// TIA Portal project "Delta_Praktika_3" (V17)

(* hardware
DEVICE "S7-1500/ET200MP station_1"  S7-1500 station
   slot 0: "Rail_0"  Rack  6ES7 590-1***0-0AA0
   slot 1: "PLC_2"  CPU 1517TF-3 PN/DP  6ES7 517-3UP00-0AB0  V2.9
      slot 3: "CPU display_1"  6ES7591-1BA00-0AA0
      slot 32768: "PROFINET interface_1"  X1
      slot 33024: "PROFINET interface_2"  X2
      slot 33280: "DP interface_1"  X3
      slot 34817: "Virtual CP interface port_1"  Virtual CP interface port  Virtual CP interface port
DEVICE "ET 200SP station_1"  ET 200SP-Station
   slot 0: "Rack_0"  Rack  6ES5 710-8MAx1
   slot 0: "et200sp"  IM 155-6 PN/2 HF  6ES7 155-6AU01-0CN0  V4.2
   slot 1: "DI 8x24VDC HF_1"  DI 8x24VDC HF  6ES7 131-6BF00-0CA0  V2.0
      slot 1: "DI 8x24VDC HF_1"  DI 8x24VDC HF
   slot 2: "DQ 8x24VDC/0.5A HF_1"  DQ 8x24VDC/0.5A HF  6ES7 132-6BF00-0CA0  V2.0
      slot 1: "DQ 8x24VDC/0.5A HF_1"  DQ 8x24VDC/0.5A HF
   slot 3: "CM 4xIO-Link_1"  CM 4xIO-Link  6ES7 137-6BD00-0BA0  V2.2
      slot 1: "CM 4xIO-Link_1"  6ES7 137-6BD00-0BA0
   slot 4: "Server module_1"  Server module  6ES7 193-6PA00-0AA0  V1.1
      slot 1: "Server module_1"  Server module
   slot 127: "BA 2xRJ45"  BA 2xRJ45  6ES7 193-6AR00-0AA0  V0.0
      slot 1: "Port_1"  X1 P1 R  6ES7 193-6AR00-0AA0  V0.0
      slot 2: "Port_2"  X1 P2 R  6ES7 193-6AR00-0AA0  V0.0
DEVICE "SINAMICS V_1"  SINAMICS V
   slot 0: "SINAMICS V90 PN Rack"  Rail  1.0
   slot 0: "a1"  V90 PN  6SL3 210-5FB10-4UFx  V1.4
      slot 1: "Drive object"  Drive Object
         slot 1: "Module access point"  Module Access Point
         slot 2: "Without PROFIsafe"  No ProfiSafe
         slot 3: "Telegram"  SIEMENS Telegramm 105
DEVICE "SINAMICS V_2"  SINAMICS V
   slot 0: "SINAMICS V90 PN Rack"  Rail  1.0
   slot 0: "a3"  V90 PN  6SL3 210-5FB10-4UFx  V1.4
      slot 1: "Drive object"  Drive Object
         slot 1: "Module access point"  Module Access Point
         slot 2: "Without PROFIsafe"  No ProfiSafe
         slot 3: "Telegram"  SIEMENS Telegramm 105
DEVICE "SINAMICS V_3"  SINAMICS V
   slot 0: "SINAMICS V90 PN Rack"  Rail  1.0
   slot 0: "a2"  V90 PN  6SL3 210-5FB10-4UFx  V1.4
      slot 1: "Drive object"  Drive Object
         slot 1: "Module access point"  Module Access Point
         slot 2: "Without PROFIsafe"  No ProfiSafe
         slot 3: "Telegram"  SIEMENS Telegramm 105
DEVICE "HMI_1"  KTP1200 Basic PN
   slot 0: "HMI_1"  KTP1200 Basic PN  6AV2 123-2MB03-0AX0  17.0.0.0
   slot 1: "HMI_RT_1"  KTP1200 Basic PN  6AV2 123-2MB03-0AX0  17.0.0.0
   slot 5: "HMI_1.IE_CP_1"  PROFINET Interface  17.0.0.0
      slot 1: "Interfaz PROFINET_1"  PROFINET Interface
         slot 1: "Port_1"  Port
*)

// ===== PLC "PLC_2"  CPU 1517TF-3 PN/DP =====
// protected blocks, not shown: "Main_Safety_RTG1", "Main_Safety_RTG1_DB"

VAR_GLOBAL   // PLC tag table "Default tag table"
   "A1_Actor_Interface_AddressIn" AT %I0.0 : "PD_TEL3_IN";
   "A1_Actor_Interface_AddressOut" AT %Q0.0 : "PD_TEL3_OUT";
   "A2_Actor_Interface_AddressIn" AT %I18.0 : "PD_TEL3_IN";
   "A2_Actor_Interface_AddressOut" AT %Q10.0 : "PD_TEL3_OUT";
   "A3_Actor_Interface_AddressIn" AT %I36.0 : "PD_TEL3_IN";
   "A3_Actor_Interface_AddressOut" AT %Q20.0 : "PD_TEL3_OUT";
   "A1_axis_Actor_Interface_AddressIn" AT %I0.0 : "PD_TEL105_IN";
   "A1_axis_Actor_Interface_AddressOut" AT %Q0.0 : "PD_TEL105_OUT";
   "a2_axis_Actor_Interface_AddressIn" AT %I20.0 : "PD_TEL105_IN";
   "a2_axis_Actor_Interface_AddressOut" AT %Q63.0 : "PD_TEL105_OUT";
   "a3_asix_Actor_Interface_AddressIn" AT %I87.0 : "PD_TEL105_IN";
   "a3_asix_Actor_Interface_AddressOut" AT %Q83.0 : "PD_TEL105_OUT";
   "Freno_a1" AT %Q30.1 : Bool;
   "marka_Freno_a1" AT %M30.1 : Bool;
   "marka_Freno_a2" AT %M30.2 : Bool;
   "Freno_a2" AT %Q30.2 : Bool;
   "Freno_a3" AT %Q30.0 : Bool;
   "marka_Freno_a3" AT %M30.0 : Bool;
   "System_Byte" AT %MB256 : Byte;
   "FirstScan" AT %M256.0 : Bool;
   "DiagStatusUpdate" AT %M256.1 : Bool;
   "AlwaysTRUE" AT %M256.2 : Bool;
   "AlwaysFALSE" AT %M256.3 : Bool;
   "Clock_Byte" AT %MB255 : Byte;
   "Clock_10Hz" AT %M255.0 : Bool;
   "Clock_5Hz" AT %M255.1 : Bool;
   "Clock_2.5Hz" AT %M255.2 : Bool;
   "Clock_2Hz" AT %M255.3 : Bool;
   "Clock_1.25Hz" AT %M255.4 : Bool;
   "Clock_1Hz" AT %M255.5 : Bool;
   "Clock_0.625Hz" AT %M255.6 : Bool;
   "Clock_0.5Hz" AT %M255.7 : Bool;
   "Tag_1" AT %M401.0 : Bool;
END_VAR

DATA_BLOCK "Power_DB"   // DB9
{ S7_Optimized_Access := 'TRUE' }
VERSION : 0.1
// stored: InstanceOfName Power
"Power"
BEGIN
END_DATA_BLOCK

DATA_BLOCK "Parametroak"   // DB11
{ S7_Optimized_Access := 'TRUE' }
VERSION : 0.1
   VAR
      Abiadura : LReal := 2.0;
      Azelerazioa : LReal := 40.0;
      Desazelerazioa : LReal := 40.0;
      Jerk : LReal := 400.0;
   END_VAR
BEGIN
END_DATA_BLOCK

DATA_BLOCK "Jog_DB"   // DB14
{ S7_Optimized_Access := 'TRUE' }
VERSION : 0.1
// stored: InstanceOfName Jog
"Jog"
BEGIN
END_DATA_BLOCK

DATA_BLOCK "Hominga_DB"   // DB18
{ S7_Optimized_Access := 'TRUE' }
VERSION : 0.1
// stored: InstanceOfName Hominga
"Hominga"
BEGIN
END_DATA_BLOCK

DATA_BLOCK "Puntuak"   // DB24
{ S7_Optimized_Access := 'TRUE' }
VERSION : 0.1
   VAR
      Puntu_abs_home : Array[1..4] of LReal;
      Puntu_abs_1 : Array[1..4] of LReal;
      Puntu_abs_2 : Array[1..4] of LReal;
      Puntu_rel_1 : Array[1..4] of LReal;
      Puntu_aux_1 : Array[1..3] of LReal;
      Puntu_zirkular_1 : Array[1..4] of LReal;
      HMI_erlatibo_lineal : Array[1..4] of LReal;
      HMI_abs_lineal : Array[1..4] of LReal;
      HMI_abs_zirkular_aux : Array[1..3] of LReal;
      HMI_abs_zirkular_endpoint : Array[1..4] of LReal;
      HMI_abs_ptp : Array[1..4] of LReal;
   END_VAR
BEGIN
   Puntu_abs_home[1] := 0.0;
   Puntu_abs_home[2] := 0.0;
   Puntu_abs_home[3] := -722.59;
   Puntu_abs_home[4] := 0.0;
   Puntu_abs_1[1] := 0.0;
   Puntu_abs_1[2] := 0.0;
   Puntu_abs_1[3] := -700.0;
   Puntu_abs_1[4] := 0.0;
   Puntu_rel_1[1] := 50.0;
   Puntu_rel_1[2] := 0.0;
   Puntu_rel_1[3] := 0.0;
   Puntu_abs_2[1] := 50.0;
   Puntu_abs_2[2] := 50.0;
   Puntu_abs_2[3] := -700.0;
   Puntu_abs_2[4] := 0.0;
   Puntu_aux_1[1] := 50.0;
   Puntu_aux_1[2] := 0.0;
   Puntu_aux_1[3] := -700.0;
   Puntu_zirkular_1[1] := 100.0;
   Puntu_zirkular_1[2] := 0.0;
   Puntu_zirkular_1[3] := -700.0;
   Puntu_zirkular_1[4] := 0.0;
END_DATA_BLOCK

DATA_BLOCK "ParametroakII"   // DB25
{ S7_Optimized_Access := 'TRUE' }
VERSION : 0.1
   VAR
      abiadura : LReal := 10.0;
      azelerazioa : LReal := 20.0;
      desazelerazioa : LReal := 20.0;
      jerk : LReal := 40.0;
   END_VAR
BEGIN
END_DATA_BLOCK

DATA_BLOCK "a1_asix"   // DB2, Motion_DB
{ S7_Optimized_Access := 'TRUE' }
AUTHOR : SIMATIC
FAMILY : MC_1500
VERSION : 6.0
// stored: InstanceOfName TO_PositioningAxis
"TO_PositioningAxis"
BEGIN
END_DATA_BLOCK

DATA_BLOCK "a2_axis"   // DB3, Motion_DB
{ S7_Optimized_Access := 'TRUE' }
AUTHOR : SIMATIC
FAMILY : MC_1500
VERSION : 6.0
// stored: InstanceOfName TO_PositioningAxis
"TO_PositioningAxis"
BEGIN
END_DATA_BLOCK

DATA_BLOCK "a3_axis"   // DB4, Motion_DB
{ S7_Optimized_Access := 'TRUE' }
AUTHOR : SIMATIC
FAMILY : MC_1500
VERSION : 6.0
// stored: InstanceOfName TO_PositioningAxis
"TO_PositioningAxis"
BEGIN
END_DATA_BLOCK

DATA_BLOCK "Delta_Robota"   // DB7, Motion_DB
{ S7_Optimized_Access := 'TRUE' }
AUTHOR : SIMATIC
FAMILY : MC_1500
VERSION : 6.0
// stored: InstanceOfName TO_Kinematics
"TO_Kinematics"
BEGIN
END_DATA_BLOCK

FUNCTION_BLOCK "Power"   // FB2, LAD
{ S7_Optimized_Access := 'TRUE' }
VERSION : 0.1
   VAR_INPUT
      Power_a1 : Bool;
      Power_a2 : Bool;
      Power_a3 : Bool;
   END_VAR
   VAR_OUTPUT
      Status_a1 : Bool;
      Status_a2 : Bool;
      Status_a3 : Bool;
      Error_a1 : Bool;
      Error_a2 : Bool;
      Error_a3 : Bool;
   END_VAR
BEGIN

REGION Network 1
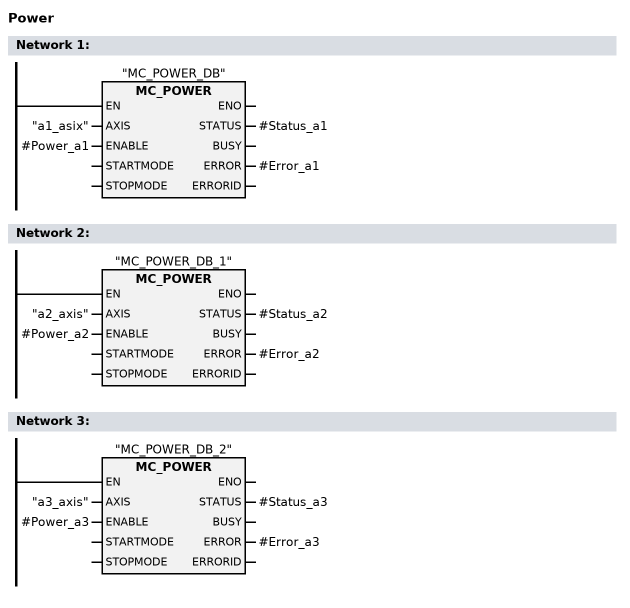
   "MC_POWER_DB"(Axis := "a1_asix", Enable := #Power_a1, Status => #Status_a1, Error => #Error_a1);   // MC_POWER
END_REGION

REGION Network 2
   "MC_POWER_DB_1"(Axis := "a2_axis", Enable := #Power_a2, Status => #Status_a2, Error => #Error_a2);   // MC_POWER
END_REGION

REGION Network 3
   "MC_POWER_DB_2"(Axis := "a3_axis", Enable := #Power_a3, Status => #Status_a3, Error => #Error_a3);   // MC_POWER
END_REGION
END_FUNCTION_BLOCK

FUNCTION_BLOCK "Jog"   // FB3, LAD
{ S7_Optimized_Access := 'TRUE' }
VERSION : 0.1
   VAR_INPUT
      "A1+" : Bool;
      "A1-" : Bool;
      "A2+" : Bool;
      "A2-" : Bool;
      "A3+" : Bool;
      "A3-" : Bool;
   END_VAR
BEGIN

REGION Network 1
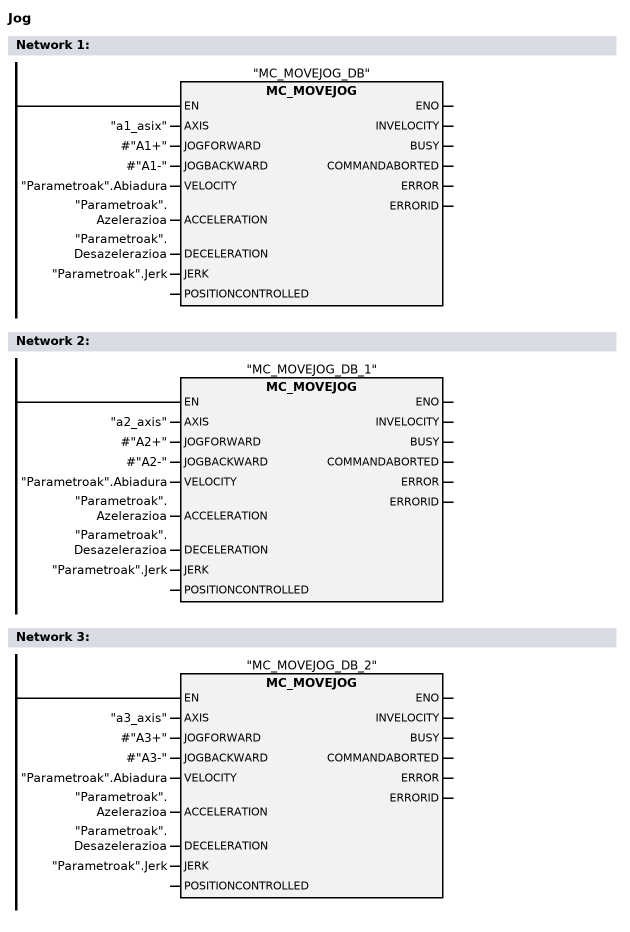
   "MC_MOVEJOG_DB"(Axis := "a1_asix",   // MC_MOVEJOG
                   JogForward := #"A1+",
                   JogBackward := #"A1-",
                   Velocity := "Parametroak".Abiadura,
                   Acceleration := "Parametroak".Azelerazioa,
                   Deceleration := "Parametroak".Desazelerazioa,
                   Jerk := "Parametroak".Jerk);
END_REGION

REGION Network 2
   "MC_MOVEJOG_DB_1"(Axis := "a2_axis",   // MC_MOVEJOG
                     JogForward := #"A2+",
                     JogBackward := #"A2-",
                     Velocity := "Parametroak".Abiadura,
                     Acceleration := "Parametroak".Azelerazioa,
                     Deceleration := "Parametroak".Desazelerazioa,
                     Jerk := "Parametroak".Jerk);
END_REGION

REGION Network 3
   "MC_MOVEJOG_DB_2"(Axis := "a3_axis",   // MC_MOVEJOG
                     JogForward := #"A3+",
                     JogBackward := #"A3-",
                     Velocity := "Parametroak".Abiadura,
                     Acceleration := "Parametroak".Azelerazioa,
                     Deceleration := "Parametroak".Desazelerazioa,
                     Jerk := "Parametroak".Jerk);
END_REGION
END_FUNCTION_BLOCK

FUNCTION_BLOCK "Hominga"   // FB4, LAD
{ S7_Optimized_Access := 'TRUE' }
VERSION : 0.1
   VAR_INPUT
      homing_a1 : Bool;
      homing_a2 : Bool;
      homing_a3 : Bool;
   END_VAR
   VAR_OUTPUT
      Done_a1 : Bool;
      Done_a2 : Bool;
      Done_a3 : Bool;
   END_VAR
BEGIN

REGION Network 1
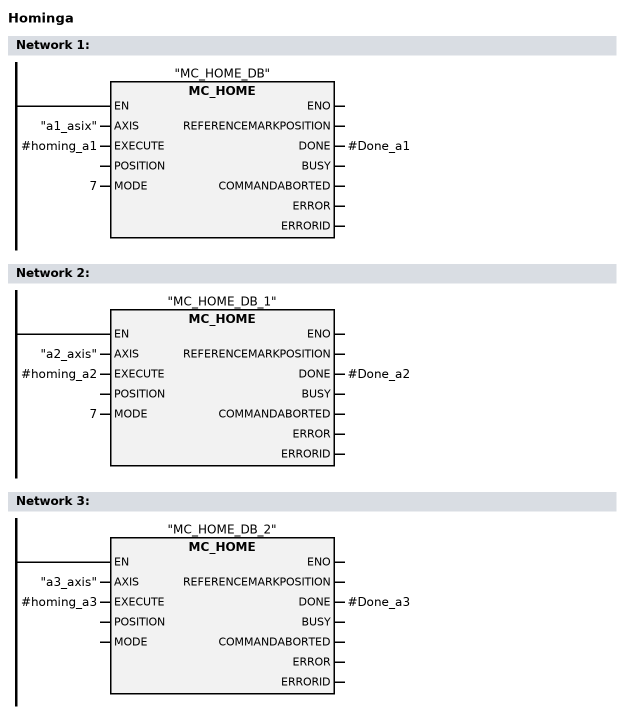
   "MC_HOME_DB"(Axis := "a1_asix", Execute := #homing_a1, Mode := 7, Done => #Done_a1);   // MC_HOME
END_REGION

REGION Network 2
   "MC_HOME_DB_1"(Axis := "a2_axis", Execute := #homing_a2, Mode := 7, Done => #Done_a2);   // MC_HOME
END_REGION

REGION Network 3
   "MC_HOME_DB_2"(Axis := "a3_axis", Execute := #homing_a3, Done => #Done_a3);   // MC_HOME
END_REGION
END_FUNCTION_BLOCK

ORGANIZATION_BLOCK "Main"   // OB1, LAD, ProgramCycle
TITLE = "Main Program Sweep (Cycle)"
{ S7_Optimized_Access := 'TRUE' }
VERSION : 0.1
   VAR_INPUT
      Initial_Call : Bool;   // Initial call of this OB
      Remanence : Bool;   // =True, if remanent data are available
   END_VAR
BEGIN

REGION Network 1
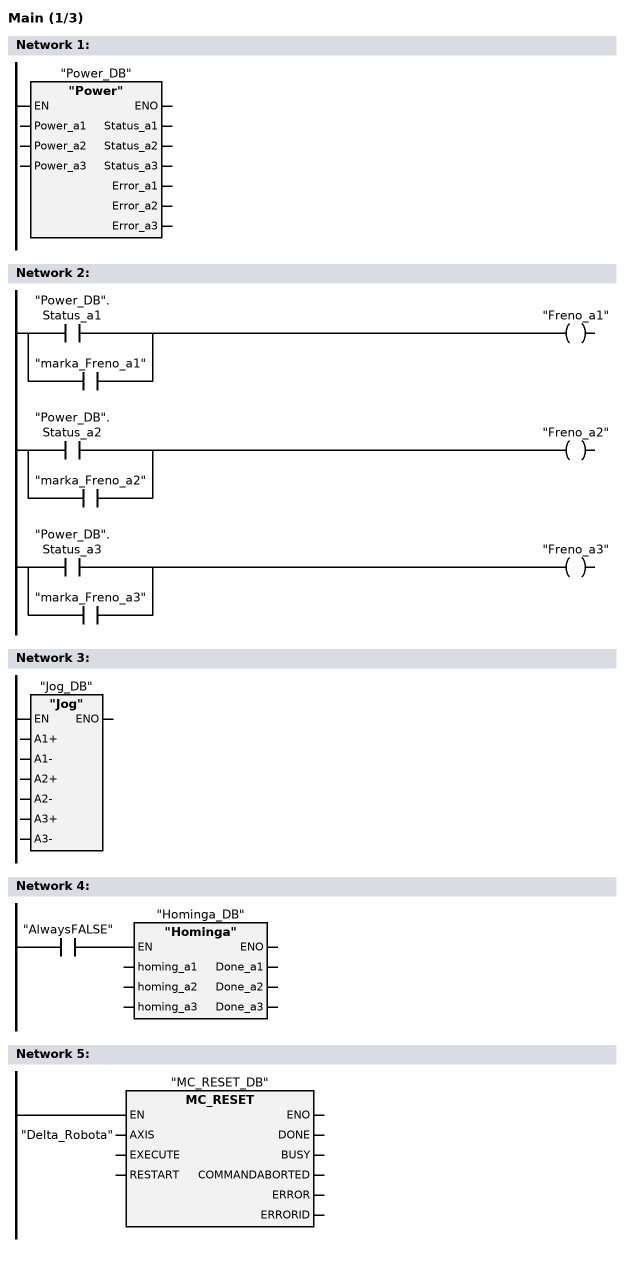
   RUNG wire#powerrail
      "Power_DB"(Power_a1 :=, Power_a2 :=, Power_a3 :=, Status_a1 =>, Status_a2 =>, Status_a3 =>, Error_a1 =>, Error_a2 =>, Error_a3 =>)
   END_RUNG
   // the same network as SCL:
   "Power_DB"();   // "Power"
END_REGION

REGION Network 2
   RUNG wire#powerrail
      Contact( "Power_DB".Status_a1 )
      wire#w1
      Coil( "Freno_a1" )
   END_RUNG
   RUNG wire#powerrail
      Contact( "marka_Freno_a1" )
   END_RUNG wire#w1
   RUNG wire#powerrail
      Contact( "Power_DB".Status_a2 )
      wire#w2
      Coil( "Freno_a2" )
   END_RUNG
   RUNG wire#powerrail
      Contact( "marka_Freno_a2" )
   END_RUNG wire#w2
   RUNG wire#powerrail
      Contact( "Power_DB".Status_a3 )
      wire#w3
      Coil( "Freno_a3" )
   END_RUNG
   RUNG wire#powerrail
      Contact( "marka_Freno_a3" )
   END_RUNG wire#w3
   // the same network as SCL:
   "Freno_a1" := "Power_DB".Status_a1 OR "marka_Freno_a1";
   "Freno_a2" := "Power_DB".Status_a2 OR "marka_Freno_a2";
   "Freno_a3" := "Power_DB".Status_a3 OR "marka_Freno_a3";
END_REGION

REGION Network 3
   RUNG wire#powerrail
      "Jog_DB"("A1+" :=, "A1-" :=, "A2+" :=, "A2-" :=, "A3+" :=, "A3-" :=)
   END_RUNG
   // the same network as SCL:
   "Jog_DB"();   // "Jog"
END_REGION

REGION Network 4
   RUNG wire#powerrail
      Contact( "AlwaysFALSE" )
      "Hominga_DB"(homing_a1 :=, homing_a2 :=, homing_a3 :=, Done_a1 =>, Done_a2 =>, Done_a3 =>)
   END_RUNG
   // the same network as SCL:
   IF "AlwaysFALSE" THEN
       "Hominga_DB"();   // "Hominga"
   END_IF;
END_REGION

REGION Network 5
   "MC_RESET_DB"(Axis := "Delta_Robota");   // MC_RESET
END_REGION

REGION Network 6
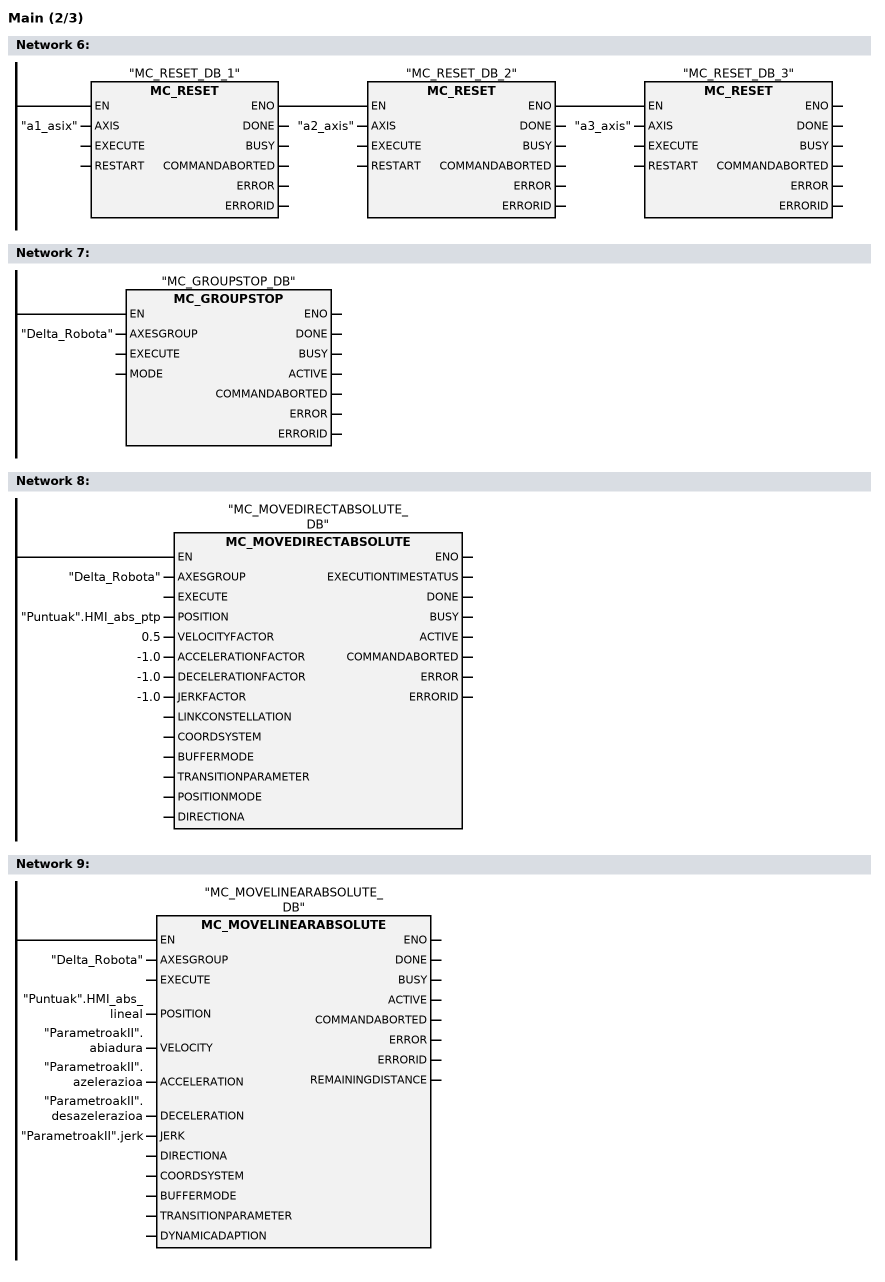
   // ENO of a box is taken as its EN; it also drops when the box reports an error
   "MC_RESET_DB_1"(Axis := "a1_asix");   // MC_RESET
   "MC_RESET_DB_2"(Axis := "a2_axis");   // MC_RESET
   "MC_RESET_DB_3"(Axis := "a3_axis");   // MC_RESET
END_REGION

REGION Network 7
   "MC_GROUPSTOP_DB"(AxesGroup := "Delta_Robota");   // MC_GROUPSTOP
END_REGION

REGION Network 8
   "MC_MOVEDIRECTABSOLUTE_DB"(AxesGroup := "Delta_Robota",   // MC_MOVEDIRECTABSOLUTE
                           Position := "Puntuak".HMI_abs_ptp,
                           VelocityFactor := 0.5,
                           AccelerationFactor := -1.0,
                           DecelerationFactor := -1.0,
                           JerkFactor := -1.0);
END_REGION

REGION Network 9
   "MC_MOVELINEARABSOLUTE_DB"(AxesGroup := "Delta_Robota",   // MC_MOVELINEARABSOLUTE
                           Position := "Puntuak".HMI_abs_lineal,
                           Velocity := "ParametroakII".abiadura,
                           Acceleration := "ParametroakII".azelerazioa,
                           Deceleration := "ParametroakII".desazelerazioa,
                           Jerk := "ParametroakII".jerk);
END_REGION

REGION Network 10
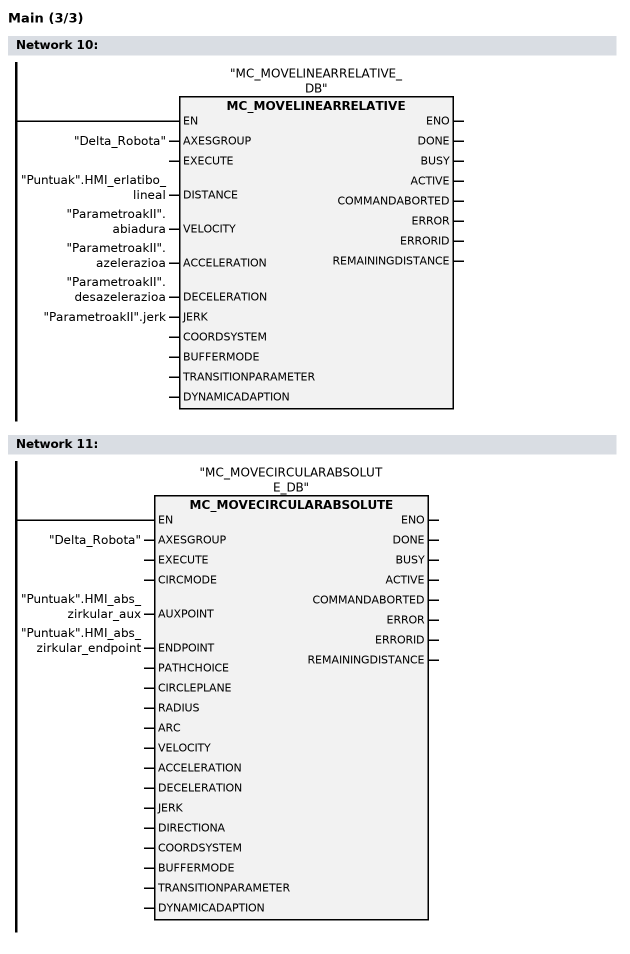
   "MC_MOVELINEARRELATIVE_DB"(AxesGroup := "Delta_Robota",   // MC_MOVELINEARRELATIVE
                           Distance := "Puntuak".HMI_erlatibo_lineal,
                           Velocity := "ParametroakII".abiadura,
                           Acceleration := "ParametroakII".azelerazioa,
                           Deceleration := "ParametroakII".desazelerazioa,
                           Jerk := "ParametroakII".jerk);
END_REGION

REGION Network 11
   "MC_MOVECIRCULARABSOLUTE_DB"(AxesGroup := "Delta_Robota",   // MC_MOVECIRCULARABSOLUTE
                           AuxPoint := "Puntuak".HMI_abs_zirkular_aux,
                           EndPoint := "Puntuak".HMI_abs_zirkular_endpoint);
END_REGION
END_ORGANIZATION_BLOCK

(* ===== HMI "HMI_RT_1" =====
system functions are stored by id; their names below are inferred from use
connection "HMI_Conexión_2": ETHERNET, SMART_S7_1500_OMS

HMI tags "Tabla de variables estándar"
   "Delta_Robota_TcpInWcs_x_Position" : LReal = PLC Delta_Robota.TcpInWcs.x.Position, 1 s
   "Power_DB_Power_a1" : Bool = PLC Power_DB.Power_a1, 1 s
   "Jog_DB_A1+" : Bool = PLC Jog_DB.A1+, 1 s
   "a1_asix_ActualPosition" : LReal = PLC a1_asix.ActualPosition, 1 s
   "Power_DB_Power_a2" : Bool = PLC Power_DB.Power_a2, 1 s
   "Power_DB_Power_a3" : Bool = PLC Power_DB.Power_a3, 1 s
   "Tag_2" : Bool = PLC marka_Freno_a1 AT %M30.1, 1 s
   "Tag_3" : Bool = PLC marka_Freno_a2 AT %M30.2, 1 s
   "Tag_6" : Bool = PLC marka_Freno_a3 AT %M30.0, 1 s
   "Jog_DB_A1-" : Bool = PLC Jog_DB.A1-, 1 s
   "Jog_DB_A2+" : Bool = PLC Jog_DB.A2+, 1 s
   "Jog_DB_A2-" : Bool = PLC Jog_DB.A2-, 1 s
   "Jog_DB_A3+" : Bool = PLC Jog_DB.A3+, 1 s
   "Jog_DB_A3-" : Bool = PLC Jog_DB.A3-, 1 s
   "Tag_1" : Bool = PLC Freno_a1 AT %Q30.1, 1 s
   "Tag_4" : Bool = PLC Freno_a2 AT %Q30.2, 1 s
   "a3_axis_ActualPosition" : LReal = PLC a3_axis.ActualPosition, 1 s
   "Tag_5" : Bool = PLC Freno_a3 AT %Q30.0, 1 s
   "Delta_Robota_TcpInWcs_y_Position" : LReal = PLC Delta_Robota.TcpInWcs.y.Position, 1 s
   "Delta_Robota_TcpInWcs_z_Position" : LReal = PLC Delta_Robota.TcpInWcs.z.Position, 1 s
   "a2_axis_ActualPosition" : LReal = PLC a2_axis.ActualPosition, 1 s
   "MC_GROUPSTOP_DB_Execute" : Bool = PLC MC_GROUPSTOP_DB.Execute, 1 s
   "MC_RESET_DB_Execute" : Bool = PLC MC_RESET_DB.Execute, 1 s
   "Puntuak_HMI_erlatibo_lineal{1}" : LReal = PLC Puntuak.HMI_erlatibo_lineal[1], 1 s
   "Puntuak_HMI_erlatibo_lineal{2}" : LReal = PLC Puntuak.HMI_erlatibo_lineal[2], 1 s
   "Puntuak_HMI_erlatibo_lineal{3}" : LReal = PLC Puntuak.HMI_erlatibo_lineal[3], 1 s
   "Puntuak_HMI_abs_lineal{1}" : LReal = PLC Puntuak.HMI_abs_lineal[1], 1 s
   "Puntuak_HMI_abs_lineal{2}" : LReal = PLC Puntuak.HMI_abs_lineal[2], 1 s
   "Puntuak_HMI_abs_lineal{3}" : LReal = PLC Puntuak.HMI_abs_lineal[3], 1 s
   "Puntuak_HMI_abs_ptp{1}" : LReal = PLC Puntuak.HMI_abs_ptp[1], 1 s
   "Puntuak_HMI_abs_ptp{2}" : LReal = PLC Puntuak.HMI_abs_ptp[2], 1 s
   "Puntuak_HMI_abs_ptp{3}" : LReal = PLC Puntuak.HMI_abs_ptp[3], 1 s
   "MC_MOVELINEARABSOLUTE_DB_Execute" : Bool = PLC MC_MOVELINEARABSOLUTE_DB.Execute, 1 s
   "MC_MOVEDIRECTABSOLUTE_DB_Execute" : Bool = PLC MC_MOVEDIRECTABSOLUTE_DB.Execute, 1 s
   "MC_MOVELINEARRELATIVE_DB_Execute" : Bool = PLC MC_MOVELINEARRELATIVE_DB.Execute, 1 s
   "Puntuak_HMI_abs_zirkular_aux{1}" : LReal = PLC Puntuak.HMI_abs_zirkular_aux[1], 1 s
   "Puntuak_HMI_abs_zirkular_aux{2}" : LReal = PLC Puntuak.HMI_abs_zirkular_aux[2], 1 s
   "Puntuak_HMI_abs_zirkular_aux{3}" : LReal = PLC Puntuak.HMI_abs_zirkular_aux[3], 1 s
   "Puntuak_HMI_abs_zirkular_endpoint{1}" : LReal = PLC Puntuak.HMI_abs_zirkular_endpoint[1], 1 s
   "Puntuak_HMI_abs_zirkular_endpoint{2}" : LReal = PLC Puntuak.HMI_abs_zirkular_endpoint[2], 1 s
   "Puntuak_HMI_abs_zirkular_endpoint{3}" : LReal = PLC Puntuak.HMI_abs_zirkular_endpoint[3], 1 s
   "MC_MOVECIRCULARABSOLUTE_DB_Execute" : Bool = PLC MC_MOVECIRCULARABSOLUTE_DB.Execute, 1 s

screen "Imagen_1" 1280x800
   Button "Botón_1" at 38,159 size 96x32; TextOff 'A1+'
      on Press: function_b14e0dd5("Jog_DB_A1+", 0)
   Button "Botón_2" at 175,159 size 96x32; TextOff 'A1-'
      on Press: function_b14e0dd5("Jog_DB_A1-", 0)
   Button "Botón_3" at 40,207 size 96x32; TextOff 'A2+'
      on Press: function_b14e0dd5("Jog_DB_A2+", 0)
   Button "Botón_4" at 175,207 size 96x32; TextOff 'A2-'
      on Press: function_b14e0dd5("Jog_DB_A2-", 0)
   Button "Botón_5" at 40,255 size 96x32; TextOff 'A3+'
      on Press: function_b14e0dd5("Jog_DB_A3+", 0)
   Button "Botón_6" at 175,255 size 96x32; TextOff 'A3-'
      on Press: function_b14e0dd5("Jog_DB_A3-", 0)
   Button "Botón_10" at 926,70 size 96x32; TextOff 'Stop'
      on Press: function_b14e0dd5("MC_GROUPSTOP_DB_Execute", 0)
   Button "Botón_11" at 1061,70 size 96x32; TextOff 'Reset'
      on Press: function_b14e0dd5("MC_RESET_DB_Execute", 0)
   TextField "Campo de texto_1" at 68,12 size 306x23; Text 'OBJETO TEKNOLOGIKOA BANAKA'
   TextField "Campo de texto_2" at 850,14 size 146x23; Text 'DELTA ROBOTA'
   Circle "Círculo_1" at 415,164 size 19x19
      Appearance <- "Tag_1"
   Circle "Círculo_2" at 415,212 size 19x19
      Appearance <- "Tag_4"
   Circle "Círculo_3" at 415,260 size 19x19
      Appearance <- "Tag_5"
   TextField "Campo de texto_3" at 144,116 size 330x23; Text 'Frenoa desaktibatuta badago berde'
   IOField "Campo ES_1" at 921,418 size 80x30; FormatPattern s999.99
      ProcessValue <- "Puntuak_HMI_abs_lineal{1}"
   IOField "Campo ES_2" at 920,452 size 81x30; FormatPattern s999.99
      ProcessValue <- "Puntuak_HMI_abs_lineal{2}"
   IOField "Campo ES_3" at 920,486 size 81x33; FormatPattern s999.99
      ProcessValue <- "Puntuak_HMI_abs_lineal{3}"
   Button "Botón_15" at 1048,454 size 96x32; TextOff 'GO!'
      on Press: function_b14e0dd5("MC_MOVELINEARABSOLUTE_DB_Execute", 0)
   TextField "Campo de texto_4" at 928,382 size 270x23; Text 'Mugimendu absoluto linearra'
   TextField "Campo de texto_5" at 1001,418 size 47x23; Text 'X'
   TextField "Campo de texto_6" at 1001,455 size 47x23; Text 'Y'
   TextField "Campo de texto_7" at 1001,492 size 47x23; Text 'Z'
   IOField "Campo ES_4" at 959,607 size 73x30; FormatPattern 99999
   IOField "Campo ES_5" at 959,641 size 73x30; FormatPattern 99999
   IOField "Campo ES_6" at 959,675 size 73x30; FormatPattern 99999
   Button "Botón_16" at 1017,715 size 96x32; TextOff 'GO!'
   TextField "Campo de texto_8" at 959,545 size 288x23; Text 'Mugimendu absoluto zirkularra'
   TextField "Campo de texto_9" at 1032,607 size 47x23; Text 'X'
   TextField "Campo de texto_10" at 1032,644 size 47x23; Text 'Y'
   TextField "Campo de texto_11" at 1032,681 size 47x23; Text 'Z'
   IOField "Campo ES_7" at 1083,608 size 73x30; FormatPattern 99999
   IOField "Campo ES_8" at 1083,642 size 73x30; FormatPattern 99999
   IOField "Campo ES_9" at 1083,676 size 73x30; FormatPattern 99999
   TextField "Campo de texto_12" at 1159,608 size 47x23; Text 'X'
   TextField "Campo de texto_13" at 1159,645 size 47x23; Text 'Y'
   TextField "Campo de texto_14" at 1159,682 size 47x23; Text 'Z'
   TextField "Campo de texto_15" at 928,575 size 135x23; Text 'Nundik pasatu'
   TextField "Campo de texto_16" at 1079,575 size 142x23; Text 'Azken posizioa'
   IOField "Campo ES_13" at 954,607 size 78x31; FormatPattern s999.99
      ProcessValue <- "Puntuak_HMI_abs_zirkular_aux{1}"
   IOField "Campo ES_14" at 954,641 size 78x30; FormatPattern s999.99
      ProcessValue <- "Puntuak_HMI_abs_zirkular_aux{2}"
   IOField "Campo ES_15" at 952,675 size 80x30; FormatPattern s999.99
      ProcessValue <- "Puntuak_HMI_abs_zirkular_aux{3}"
   Button "Botón_18" at 1017,715 size 96x32; TextOff 'GO!'
      on Press: function_b14e0dd5("MC_MOVECIRCULARABSOLUTE_DB_Execute", 0)
   TextField "Campo de texto_21" at 959,545 size 288x23; Text 'Mugimendu absoluto zirkularra'
   TextField "Campo de texto_22" at 1032,607 size 47x23; Text 'X'
   TextField "Campo de texto_23" at 1032,644 size 47x23; Text 'Y'
   TextField "Campo de texto_24" at 1032,681 size 47x23; Text 'Z'
   IOField "Campo ES_16" at 1077,608 size 79x30; FormatPattern s999.99
      ProcessValue <- "Puntuak_HMI_abs_zirkular_endpoint{1}"
   IOField "Campo ES_17" at 1078,642 size 78x30; FormatPattern s999.99
      ProcessValue <- "Puntuak_HMI_abs_zirkular_endpoint{2}"
   IOField "Campo ES_18" at 1078,676 size 78x30; FormatPattern s999.99
      ProcessValue <- "Puntuak_HMI_abs_zirkular_endpoint{3}"
   TextField "Campo de texto_25" at 1159,608 size 47x23; Text 'X'
   TextField "Campo de texto_26" at 1159,645 size 47x23; Text 'Y'
   TextField "Campo de texto_27" at 1159,682 size 47x23; Text 'Z'
   TextField "Campo de texto_28" at 928,575 size 135x23; Text 'Nundik pasatu'
   TextField "Campo de texto_29" at 1079,575 size 142x23; Text 'Azken posizioa'
   IOField "Campo ES_10" at 40,390 size 96x32; FormatPattern s99.999
      ProcessValue <- "a1_asix_ActualPosition"
   IOField "Campo ES_11" at 166,388 size 96x32; FormatPattern s99.999
      ProcessValue <- "a2_axis_ActualPosition"
   IOField "Campo ES_12" at 308,388 size 96x32; FormatPattern s99.999
      ProcessValue <- "a3_axis_ActualPosition"
   TextField "Campo de texto_17" at 68,352 size 46x25; Text 'A1'
   TextField "Campo de texto_18" at 198,352 size 46x25; Text 'A2'
   TextField "Campo de texto_19" at 328,352 size 46x25; Text 'A3'
   IOField "Campo ES_19" at 549,418 size 86x33; FormatPattern s999.99
      ProcessValue <- "Puntuak_HMI_erlatibo_lineal{1}"
   IOField "Campo ES_20" at 550,452 size 85x31; FormatPattern s999.99
      ProcessValue <- "Puntuak_HMI_erlatibo_lineal{2}"
   IOField "Campo ES_21" at 550,486 size 85x30; FormatPattern s999.99
      ProcessValue <- "Puntuak_HMI_erlatibo_lineal{3}"
   Button "Botón_17" at 682,454 size 96x32; TextOff 'GO!'
      on Press: function_b14e0dd5("MC_MOVELINEARRELATIVE_DB_Execute", 0)
   TextField "Campo de texto_20" at 562,382 size 264x23; Text 'Mugimendu erlatibo linearra'
   TextField "Campo de texto_30" at 635,418 size 47x23; Text 'X'
   TextField "Campo de texto_31" at 635,455 size 47x23; Text 'Y'
   TextField "Campo de texto_32" at 635,492 size 47x23; Text 'Z'
   IOField "Campo ES_25" at 594,613 size 73x30; FormatPattern 99999
   IOField "Campo ES_26" at 594,647 size 73x30; FormatPattern 99999
   IOField "Campo ES_27" at 594,681 size 73x30; FormatPattern 99999
   TextField "Campo de texto_37" at 682,618 size 47x23; Text 'X'
   TextField "Campo de texto_38" at 682,655 size 47x23; Text 'Y'
   TextField "Campo de texto_39" at 682,692 size 47x23; Text 'Z'
   Button "Botón_20" at 713,649 size 96x32; TextOff 'GO!'
      on Press: function_b14e0dd5("MC_MOVEDIRECTABSOLUTE_DB_Execute", 0)
   IOField "Campo ES_31" at 585,613 size 82x31; FormatPattern s999.99
      ProcessValue <- "Puntuak_HMI_abs_ptp{1}"
   IOField "Campo ES_32" at 584,647 size 83x31; FormatPattern s999.99
      ProcessValue <- "Puntuak_HMI_abs_ptp{2}"
   IOField "Campo ES_33" at 584,681 size 83x29; FormatPattern s999.99
      ProcessValue <- "Puntuak_HMI_abs_ptp{3}"
   TextField "Campo de texto_46" at 682,618 size 47x23; Text 'X'
   TextField "Campo de texto_47" at 682,655 size 47x23; Text 'Y'
   TextField "Campo de texto_48" at 682,692 size 47x23; Text 'Z'
   TextField "Campo de texto_42" at 581,326 size 254x25; Text 'MUGIMENDU ERLATIBOAK'
   TextField "Campo de texto_51" at 603,540 size 261x25; Text 'MUGIMENDU ABSOLUTOAK'
   IOField "Campo ES_34" at 532,119 size 96x32; FormatPattern s999.999
      ProcessValue <- "Delta_Robota_TcpInWcs_x_Position"
   IOField "Campo ES_35" at 532,179 size 96x32; FormatPattern s999.999
      ProcessValue <- "Delta_Robota_TcpInWcs_y_Position"
   IOField "Campo ES_36" at 532,239 size 96x32; FormatPattern s999.999
      ProcessValue <- "Delta_Robota_TcpInWcs_z_Position"
   TextField "Campo de texto_52" at 635,123 size 46x25; Text 'X'
   TextField "Campo de texto_53" at 633,181 size 46x25; Text 'Y'
   TextField "Campo de texto_54" at 636,239 size 46x25; Text 'Z'
   TextField "Campo de texto_55" at 506,79 size 284x25; Text 'MOMENTUKO X Y Z POSIZIOA'
   TextField "Campo de texto_56" at 14,304 size 448x25; Text 'MOMENTUKO ARDATZEN POSIZIOA GRADUTAN'
   Button "Botón_21" at 888,150 size 298x100; TextOff 'Pick & Place MARTXA'
   Switch "Interruptor_1" at 52,70 size 64x32; CaptionText 'Switch'; TextOff 'OFF'; TextOn 'ON'
      on SwitchOn: SetBit("Power_DB_Power_a1")
      on SwitchOff: ResetBit("Power_DB_Power_a1")
   TextField "Campo de texto_57" at 52,45 size 87x25; Text 'Power A1'
   Switch "Interruptor_2" at 187,70 size 64x32; TextOn 'ON'; CaptionText 'Switch'; TextOff 'OFF'
      on SwitchOn: SetBit("Power_DB_Power_a2")
      on SwitchOff: ResetBit("Power_DB_Power_a2")
   TextField "Campo de texto_58" at 187,45 size 87x25; Text 'Power A2'
   Switch "Interruptor_3" at 322,70 size 64x32; TextOn 'ON'; CaptionText 'Switch'; TextOff 'OFF'
      on SwitchOff: ResetBit("Power_DB_Power_a3")
      on SwitchOn: SetBit("Power_DB_Power_a3")
   TextField "Campo de texto_59" at 322,45 size 87x25; Text 'Power A3'
   Switch "Interruptor_4" at 322,159 size 64x32; TextOn 'ON'; CaptionText 'Switch'; TextOff 'OFF'
      on SwitchOff: ResetBit("Tag_2")
      on SwitchOn: SetBit("Tag_2")
   Switch "Interruptor_5" at 322,207 size 64x32; TextOn 'ON'; CaptionText 'Switch'; TextOff 'OFF'
      on SwitchOff: ResetBit("Tag_3")
      on SwitchOn: SetBit("Tag_3")
   Switch "Interruptor_6" at 322,256 size 64x32; TextOn 'ON'; CaptionText 'Switch'; TextOff 'OFF'
      on SwitchOn: SetBit("Tag_6")
      on SwitchOff: ResetBit("Tag_6")
   TextField "Campo de texto_60" at 315,135 size 82x25; Text 'Freno A1'
   TextField "Campo de texto_61" at 315,187 size 82x25; Text 'Freno A2'
   TextField "Campo de texto_62" at 315,235 size 82x25; Text 'Freno A3'
   TextField "Campo de texto_33" at 952,334 size 241x25; Text 'MUGIMENDU ABSOLUTOAK'
   TextField "Campo de texto_40" at 569,568 size 290x23; Text 'Mugimendu absoluto point to point'
*)